(* Logix 5000 project; controller PLC_MCC1300_75F1 vendor 1 type 14 code 166 rev 32.11; software revision 32.04; part 44 of 83 *)
(* tags used below, declared in another part *)
   CONST_tPlant : UDT_PLANT_CONSTANTS;
   GP_OB_InitializeMain : GP_OB_Initialize;
   GP_PosWindow : GP_PosWindow;
   GP_TrackingSearchPlate : GP_TrackingSearchPlate;
   M307ASpeedUp : MAC_SpeedUp;
   M307ASpeedUp_ALM : MAC_SpeedUp_ALM;
   M30xTrimDeck : MAC_TrimmingDeck[5];
   M30xTrimDeck_ALM : MAC_TrimmingDeck_ALM[5];
   M30xTrimDeck_HMR : MAC_TrimmingDeck_HMR[5];
   TMP_d : DINT;
   TMP_dIndex : DINT;
   TMP_dIndexMotor : DINT;
   TMP_dLineSpeed : DINT;
   TMP_r : REAL;
   TMP_x : BOOL;
   xAlwaysOFF : BOOL;
   xDebugOFF : BOOL;
   Z200_SnapDataEth : UDT_ConvoyCap_ZC[2];
   Z300_BufferPlate : UDT_LINE_BUFFER_PLATE;
   Z300_Conveyor : UDT_StandConv[29];
   Z300_LineTracking : UDT_LINE_TRACKING;
   Z301 : MAC_Zone_ML;
   Z301_HMR : MAC_Zone_ML_HMR;
   Z301_HMW : MAC_Zone_ML_HMW;
(* MainProgram, continued *)

ROUTINE M307ASpeedUp_Faults   (* ladder *)
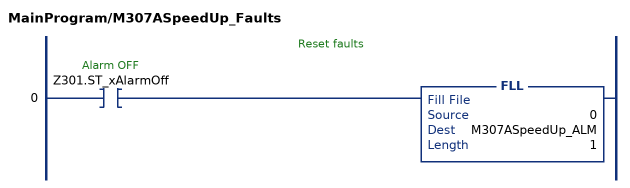
   // Reset faults
   0: XIC(Z301.ST_xAlarmOff)FLL(0,M307ASpeedUp_ALM,1);
END_ROUTINE

ROUTINE M307ASpeedUp_Logic   (* ladder *)
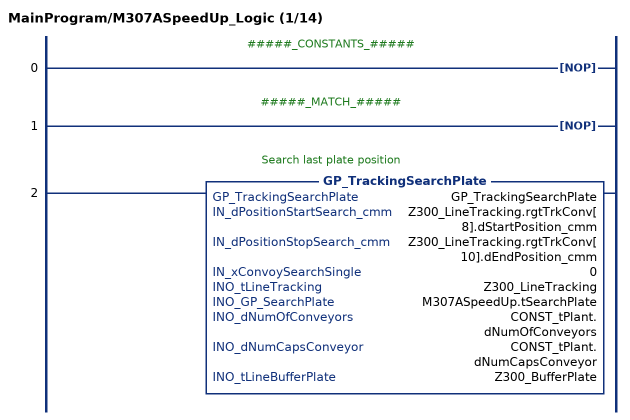
   // #####_CONSTANTS_#####
   0: NOP();
   // #####_MATCH_#####
   1: NOP();
   // Search last plate position
   2: GP_TrackingSearchPlate(GP_TrackingSearchPlate,Z300_LineTracking.rgtTrkConv[8].dStartPosition_cmm,Z300_LineTracking.rgtTrkConv[10].dEndPosition_cmm,0,Z300_LineTracking,M307ASpeedUp.tSearchPlate,CONST_tPlant.dNumOfConveyors,CONST_tPlant.dNumCapsConveyor,Z300_BufferPlate);
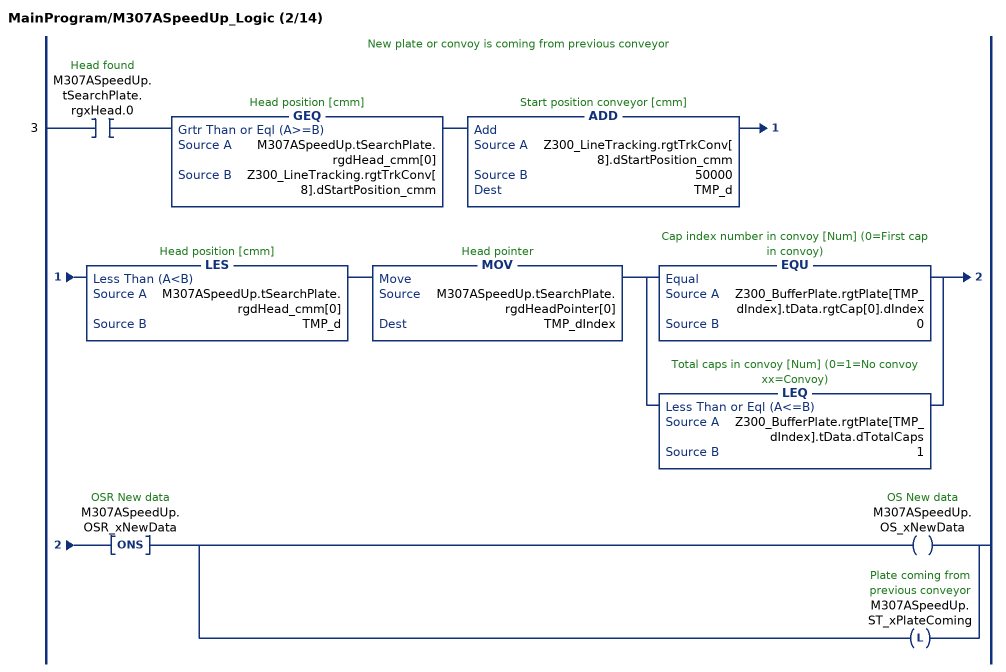
   // New plate or convoy is coming from previous conveyor
   3: XIC(M307ASpeedUp.tSearchPlate.rgxHead.0)GEQ(M307ASpeedUp.tSearchPlate.rgdHead_cmm[0],Z300_LineTracking.rgtTrkConv[8].dStartPosition_cmm)ADD(Z300_LineTracking.rgtTrkConv[8].dStartPosition_cmm,50000,TMP_d)LES(M307ASpeedUp.tSearchPlate.rgdHead_cmm[0],TMP_d)MOV(M307ASpeedUp.tSearchPlate.rgdHeadPointer[0],TMP_dIndex)[EQU(Z300_BufferPlate.rgtPlate[TMP_dIndex].tData.rgtCap[0].dIndex,0) ,LEQ(Z300_BufferPlate.rgtPlate[TMP_dIndex].tData.dTotalCaps,1) ]ONS(M307ASpeedUp.OSR_xNewData)[OTE(M307ASpeedUp.OS_xNewData) ,OTL(M307ASpeedUp.ST_xPlateComing) ];
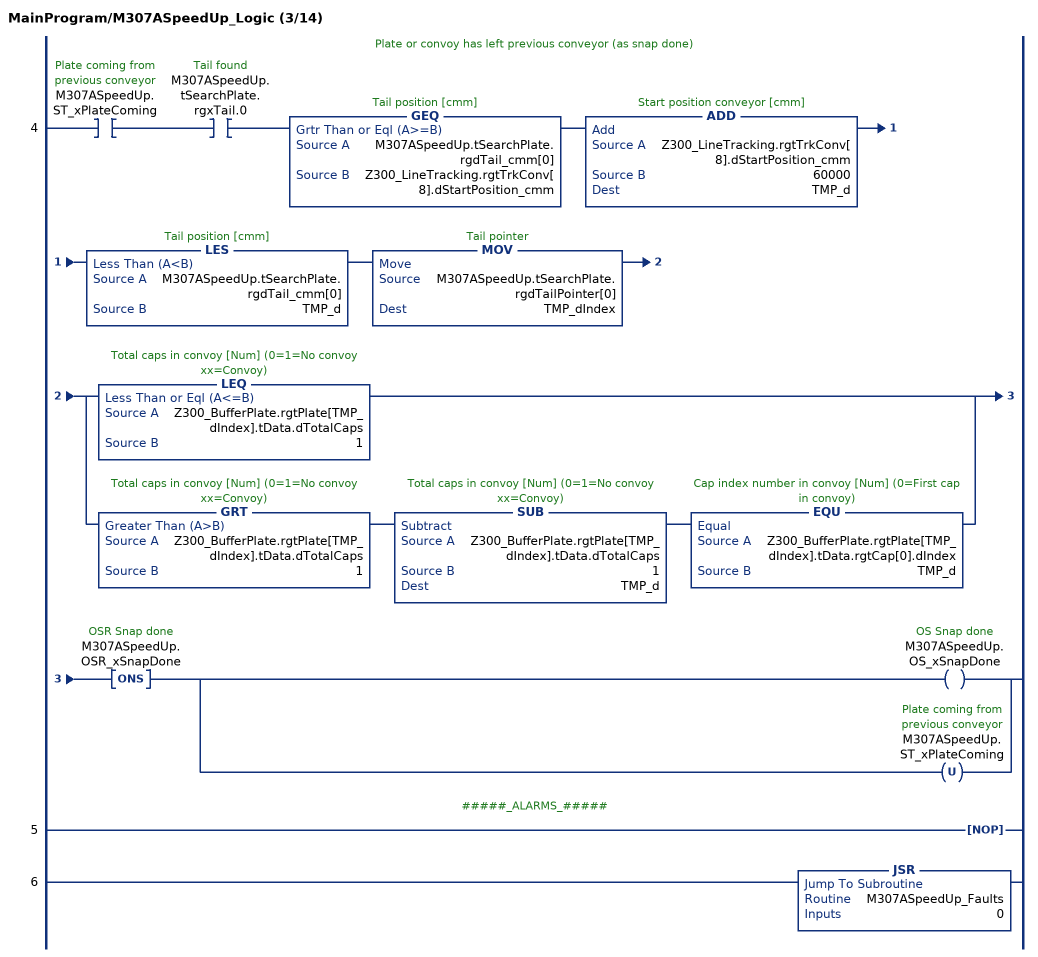
   // Plate or convoy has left previous conveyor (as snap done)
   4: XIC(M307ASpeedUp.ST_xPlateComing)XIC(M307ASpeedUp.tSearchPlate.rgxTail.0)GEQ(M307ASpeedUp.tSearchPlate.rgdTail_cmm[0],Z300_LineTracking.rgtTrkConv[8].dStartPosition_cmm)ADD(Z300_LineTracking.rgtTrkConv[8].dStartPosition_cmm,60000,TMP_d)LES(M307ASpeedUp.tSearchPlate.rgdTail_cmm[0],TMP_d)MOV(M307ASpeedUp.tSearchPlate.rgdTailPointer[0],TMP_dIndex)[LEQ(Z300_BufferPlate.rgtPlate[TMP_dIndex].tData.dTotalCaps,1) ,GRT(Z300_BufferPlate.rgtPlate[TMP_dIndex].tData.dTotalCaps,1) SUB(Z300_BufferPlate.rgtPlate[TMP_dIndex].tData.dTotalCaps,1,TMP_d) EQU(Z300_BufferPlate.rgtPlate[TMP_dIndex].tData.rgtCap[0].dIndex,TMP_d) ]ONS(M307ASpeedUp.OSR_xSnapDone)[OTE(M307ASpeedUp.OS_xSnapDone) ,OTU(M307ASpeedUp.ST_xPlateComing) ];
   // #####_ALARMS_#####
   5: NOP();
   6: JSR(M307ASpeedUp_Faults,0);
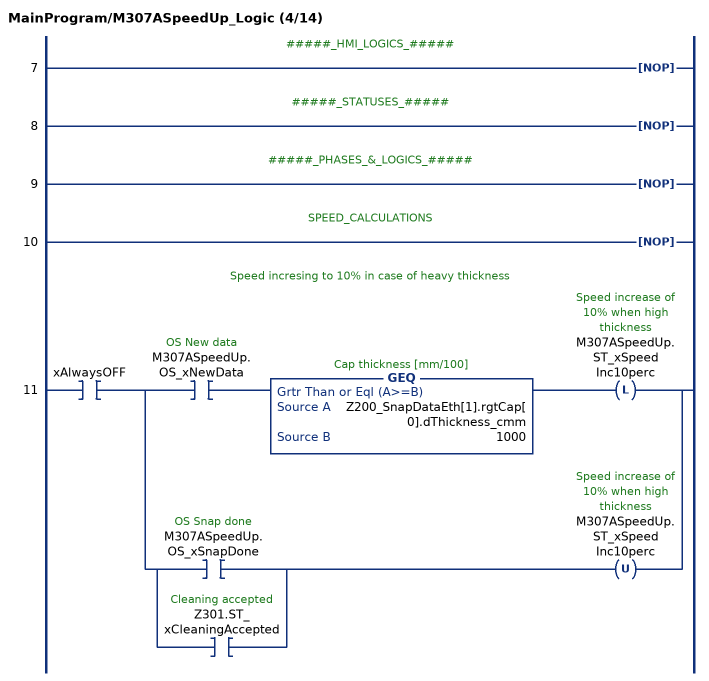
   // #####_HMI_LOGICS_#####
   7: NOP();
   // #####_STATUSES_#####
   8: NOP();
   // #####_PHASES_&_LOGICS_#####
   9: NOP();
   // SPEED_CALCULATIONS
   10: NOP();
   // Speed incresing to 10% in case of heavy thickness
   11: XIC(xAlwaysOFF)[XIC(M307ASpeedUp.OS_xNewData) GEQ(Z200_SnapDataEth[1].rgtCap[0].dThickness_cmm,1000) OTL(M307ASpeedUp.ST_xSpeedInc10perc) ,[XIC(M307ASpeedUp.OS_xSnapDone) ,XIC(Z301.ST_xCleaningAccepted) ] OTU(M307ASpeedUp.ST_xSpeedInc10perc) ];
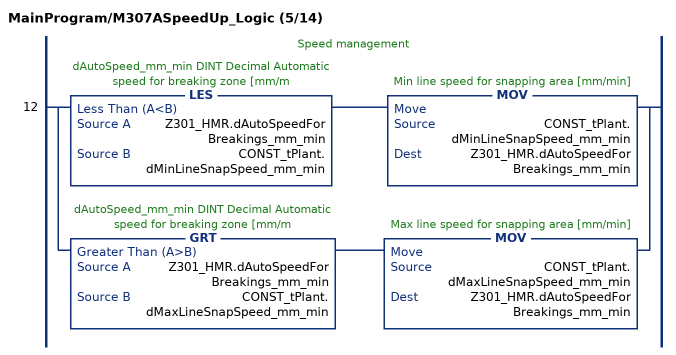
   // Speed management
   12: [LES(Z301_HMR.dAutoSpeedForBreakings_mm_min,CONST_tPlant.dMinLineSnapSpeed_mm_min) MOV(CONST_tPlant.dMinLineSnapSpeed_mm_min,Z301_HMR.dAutoSpeedForBreakings_mm_min) ,GRT(Z301_HMR.dAutoSpeedForBreakings_mm_min,CONST_tPlant.dMaxLineSnapSpeed_mm_min) MOV(CONST_tPlant.dMaxLineSnapSpeed_mm_min,Z301_HMR.dAutoSpeedForBreakings_mm_min) ];
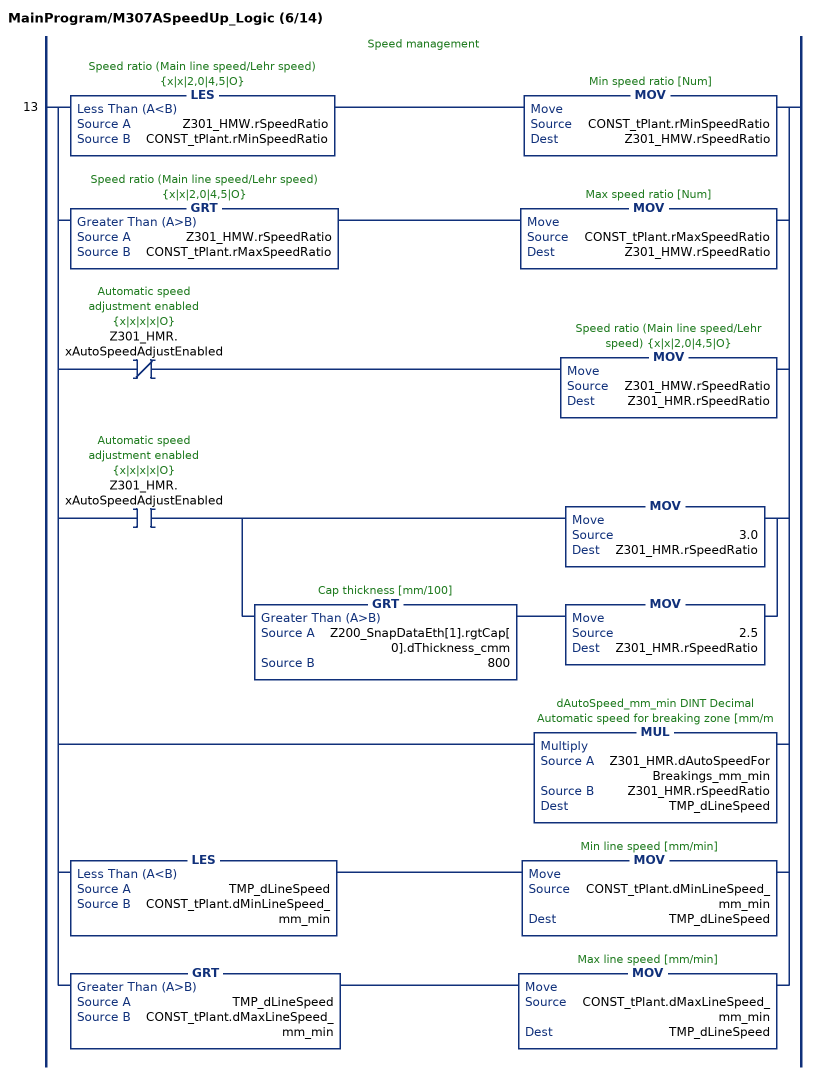
   // Speed management
   13: [LES(Z301_HMW.rSpeedRatio,CONST_tPlant.rMinSpeedRatio) MOV(CONST_tPlant.rMinSpeedRatio,Z301_HMW.rSpeedRatio) ,GRT(Z301_HMW.rSpeedRatio,CONST_tPlant.rMaxSpeedRatio) MOV(CONST_tPlant.rMaxSpeedRatio,Z301_HMW.rSpeedRatio) ,XIO(Z301_HMR.xAutoSpeedAdjustEnabled) MOV(Z301_HMW.rSpeedRatio,Z301_HMR.rSpeedRatio) ,XIC(Z301_HMR.xAutoSpeedAdjustEnabled) [MOV(3.0,Z301_HMR.rSpeedRatio) ,GRT(Z200_SnapDataEth[1].rgtCap[0].dThickness_cmm,800) MOV(2.5,Z301_HMR.rSpeedRatio) ] ,MUL(Z301_HMR.dAutoSpeedForBreakings_mm_min,Z301_HMR.rSpeedRatio,TMP_dLineSpeed) ,LES(TMP_dLineSpeed,CONST_tPlant.dMinLineSpeed_mm_min) MOV(CONST_tPlant.dMinLineSpeed_mm_min,TMP_dLineSpeed) ,GRT(TMP_dLineSpeed,CONST_tPlant.dMaxLineSpeed_mm_min) MOV(CONST_tPlant.dMaxLineSpeed_mm_min,TMP_dLineSpeed) ];
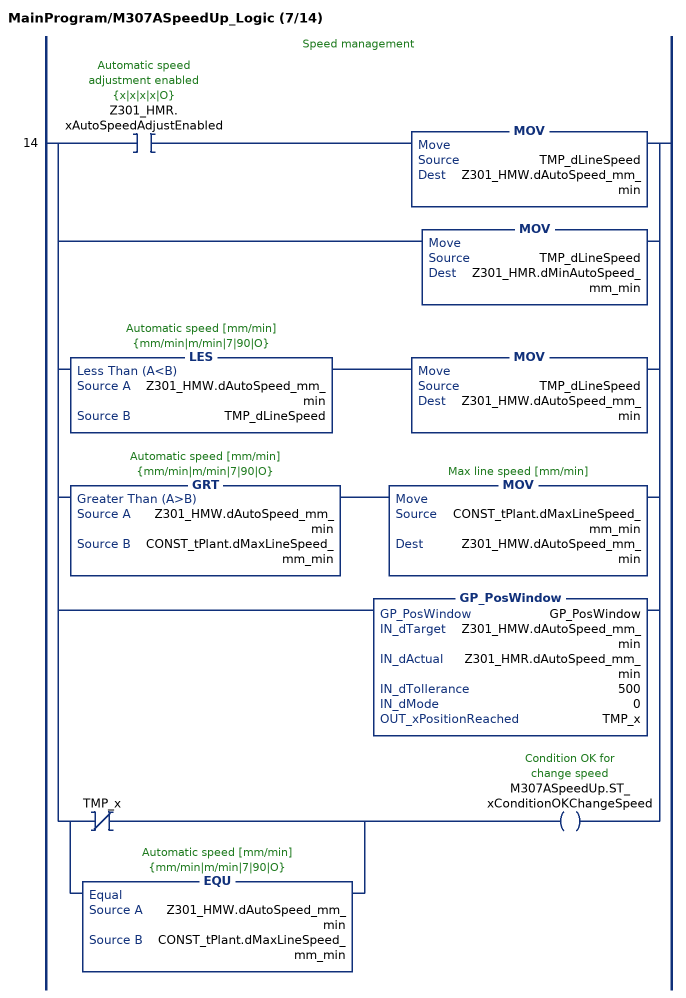
   // Speed management
   14: [XIC(Z301_HMR.xAutoSpeedAdjustEnabled) MOV(TMP_dLineSpeed,Z301_HMW.dAutoSpeed_mm_min) ,MOV(TMP_dLineSpeed,Z301_HMR.dMinAutoSpeed_mm_min) ,LES(Z301_HMW.dAutoSpeed_mm_min,TMP_dLineSpeed) MOV(TMP_dLineSpeed,Z301_HMW.dAutoSpeed_mm_min) ,GRT(Z301_HMW.dAutoSpeed_mm_min,CONST_tPlant.dMaxLineSpeed_mm_min) MOV(CONST_tPlant.dMaxLineSpeed_mm_min,Z301_HMW.dAutoSpeed_mm_min) ,[GP_PosWindow(GP_PosWindow,Z301_HMW.dAutoSpeed_mm_min,Z301_HMR.dAutoSpeed_mm_min,500,0,TMP_x) ,[XIO(TMP_x) ,EQU(Z301_HMW.dAutoSpeed_mm_min,CONST_tPlant.dMaxLineSpeed_mm_min) ] OTE(M307ASpeedUp.ST_xConditionOKChangeSpeed) ] ];
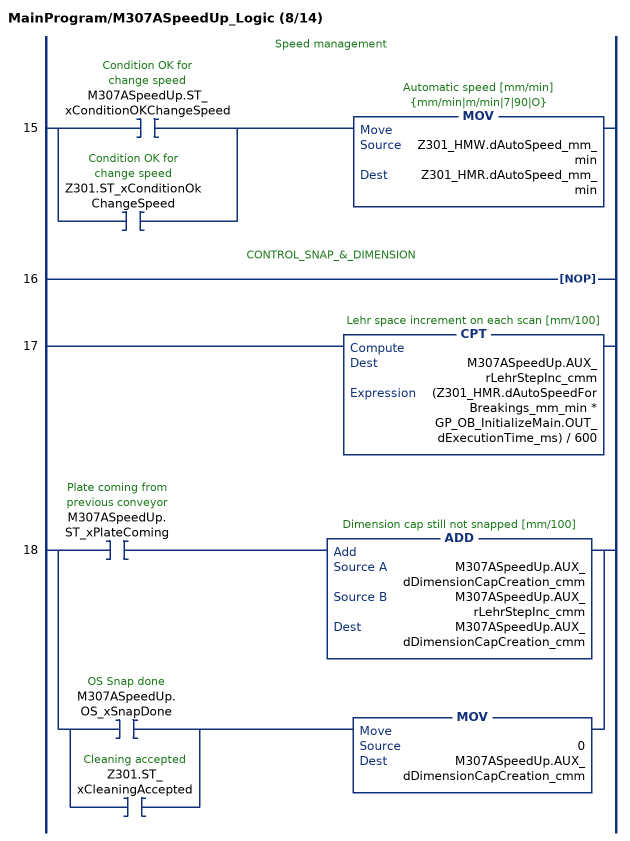
   // Speed management
   15: [XIC(M307ASpeedUp.ST_xConditionOKChangeSpeed) ,XIC(Z301.ST_xConditionOkChangeSpeed) ]MOV(Z301_HMW.dAutoSpeed_mm_min,Z301_HMR.dAutoSpeed_mm_min);
   // CONTROL_SNAP_&_DIMENSION
   16: NOP();
   17: CPT(M307ASpeedUp.AUX_rLehrStepInc_cmm,(Z301_HMR.dAutoSpeedForBreakings_mm_min * GP_OB_InitializeMain.OUT_dExecutionTime_ms) / 600);
   18: [XIC(M307ASpeedUp.ST_xPlateComing) ADD(M307ASpeedUp.AUX_dDimensionCapCreation_cmm,M307ASpeedUp.AUX_rLehrStepInc_cmm,M307ASpeedUp.AUX_dDimensionCapCreation_cmm) ,[XIC(M307ASpeedUp.OS_xSnapDone) ,XIC(Z301.ST_xCleaningAccepted) ] MOV(0,M307ASpeedUp.AUX_dDimensionCapCreation_cmm) ];
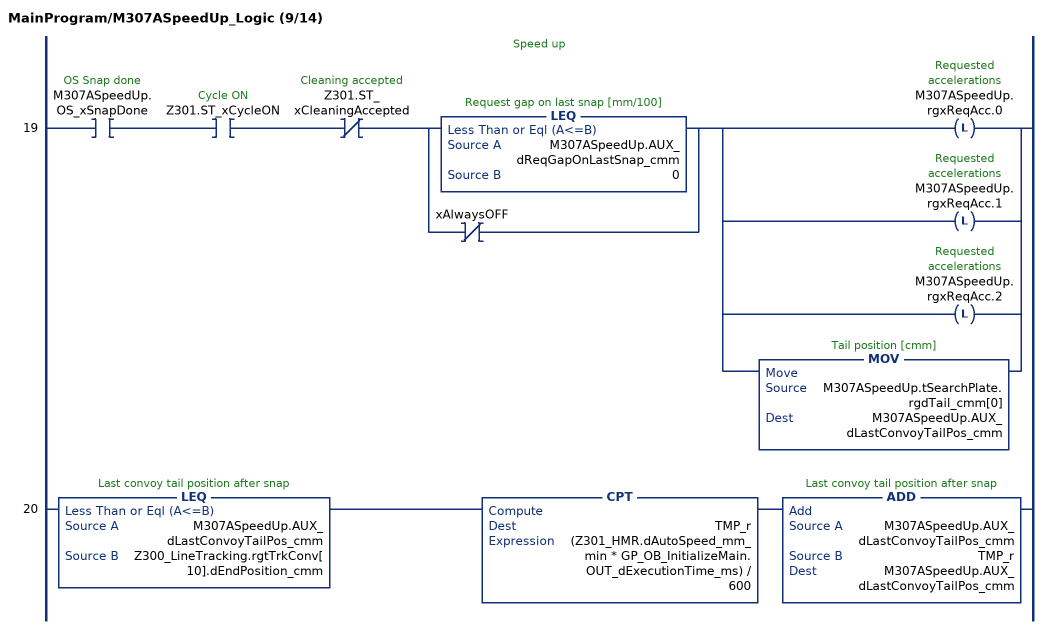
   // Speed up
   19: XIC(M307ASpeedUp.OS_xSnapDone)XIC(Z301.ST_xCycleON)XIO(Z301.ST_xCleaningAccepted)[LEQ(M307ASpeedUp.AUX_dReqGapOnLastSnap_cmm,0) ,XIO(xAlwaysOFF) ][OTL(M307ASpeedUp.rgxReqAcc.0) ,OTL(M307ASpeedUp.rgxReqAcc.1) ,OTL(M307ASpeedUp.rgxReqAcc.2) ,MOV(M307ASpeedUp.tSearchPlate.rgdTail_cmm[0],M307ASpeedUp.AUX_dLastConvoyTailPos_cmm) ];
   20: LEQ(M307ASpeedUp.AUX_dLastConvoyTailPos_cmm,Z300_LineTracking.rgtTrkConv[10].dEndPosition_cmm)CPT(TMP_r,(Z301_HMR.dAutoSpeed_mm_min * GP_OB_InitializeMain.OUT_dExecutionTime_ms) / 600)ADD(M307ASpeedUp.AUX_dLastConvoyTailPos_cmm,TMP_r,M307ASpeedUp.AUX_dLastConvoyTailPos_cmm);
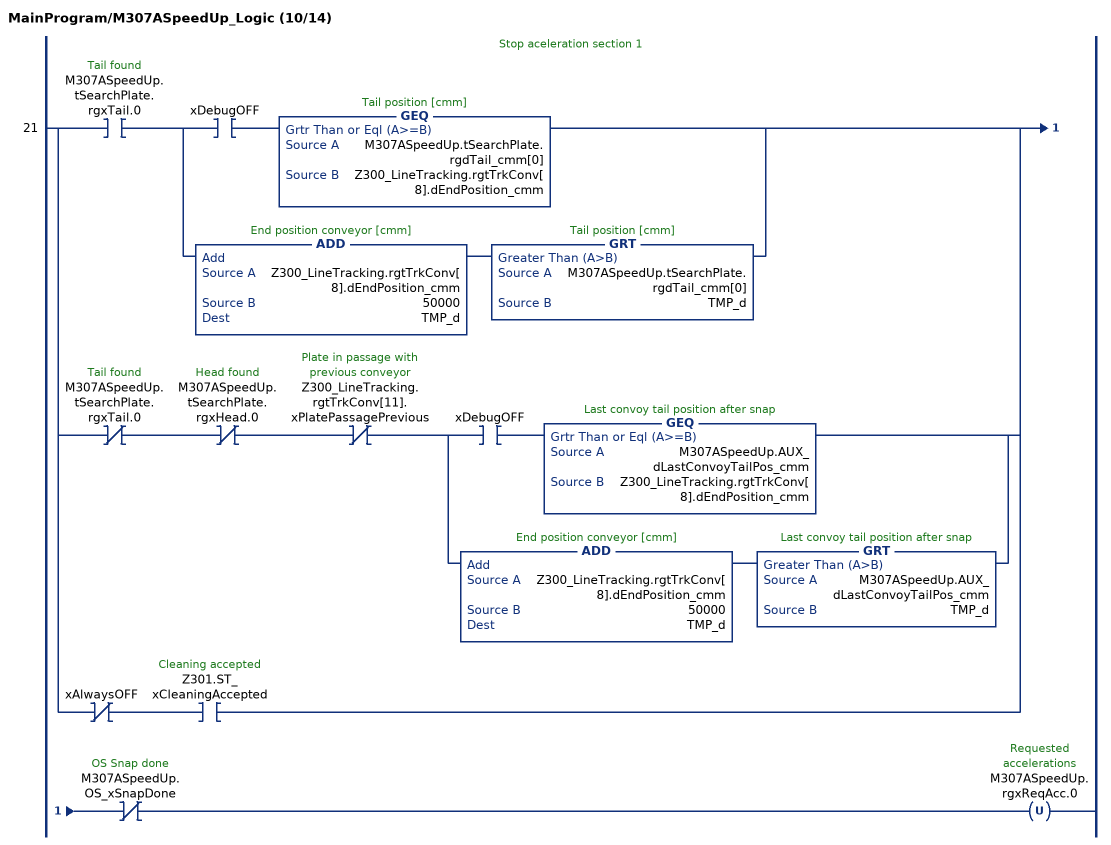
   // Stop aceleration section 1
   21: [XIC(M307ASpeedUp.tSearchPlate.rgxTail.0) [XIC(xDebugOFF) GEQ(M307ASpeedUp.tSearchPlate.rgdTail_cmm[0],Z300_LineTracking.rgtTrkConv[8].dEndPosition_cmm) ,ADD(Z300_LineTracking.rgtTrkConv[8].dEndPosition_cmm,50000,TMP_d) GRT(M307ASpeedUp.tSearchPlate.rgdTail_cmm[0],TMP_d) ] ,XIO(M307ASpeedUp.tSearchPlate.rgxTail.0) XIO(M307ASpeedUp.tSearchPlate.rgxHead.0) XIO(Z300_LineTracking.rgtTrkConv[11].xPlatePassagePrevious) [XIC(xDebugOFF) GEQ(M307ASpeedUp.AUX_dLastConvoyTailPos_cmm,Z300_LineTracking.rgtTrkConv[8].dEndPosition_cmm) ,ADD(Z300_LineTracking.rgtTrkConv[8].dEndPosition_cmm,50000,TMP_d) GRT(M307ASpeedUp.AUX_dLastConvoyTailPos_cmm,TMP_d) ] ,XIO(xAlwaysOFF) XIC(Z301.ST_xCleaningAccepted) ]XIO(M307ASpeedUp.OS_xSnapDone)OTU(M307ASpeedUp.rgxReqAcc.0);
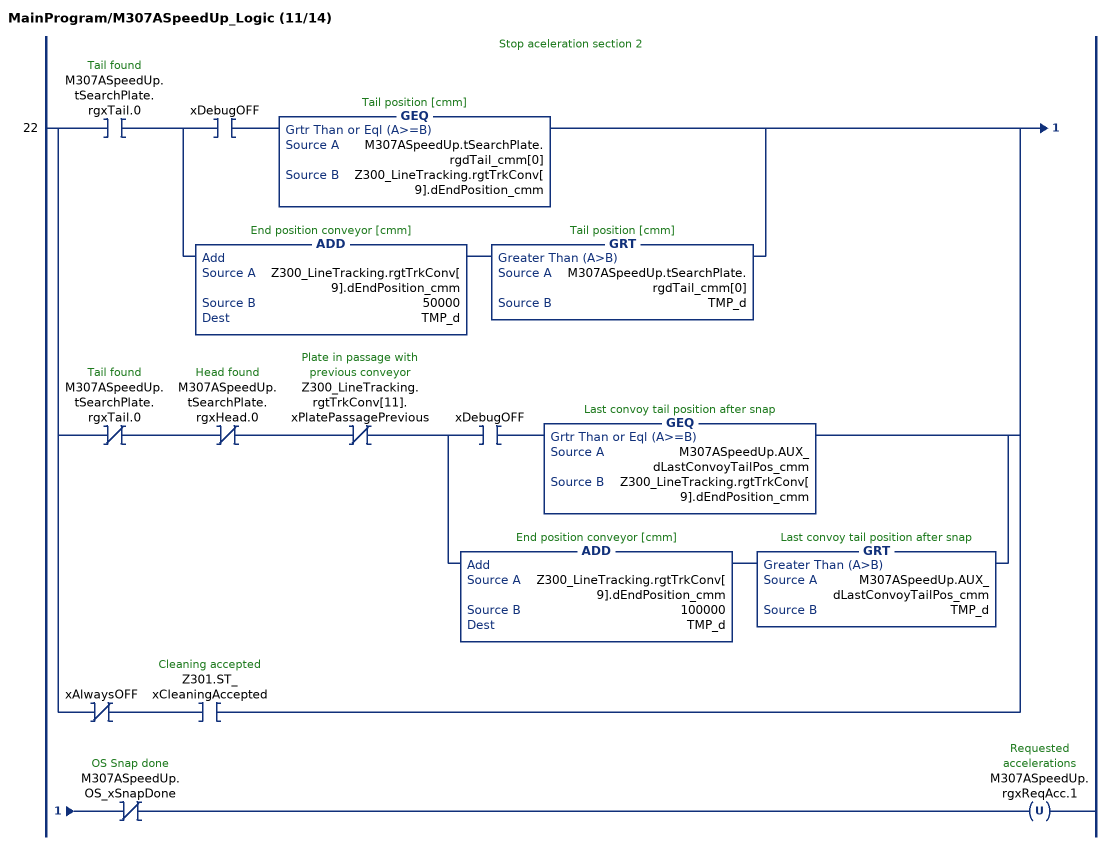
   // Stop aceleration section 2
   22: [XIC(M307ASpeedUp.tSearchPlate.rgxTail.0) [XIC(xDebugOFF) GEQ(M307ASpeedUp.tSearchPlate.rgdTail_cmm[0],Z300_LineTracking.rgtTrkConv[9].dEndPosition_cmm) ,ADD(Z300_LineTracking.rgtTrkConv[9].dEndPosition_cmm,50000,TMP_d) GRT(M307ASpeedUp.tSearchPlate.rgdTail_cmm[0],TMP_d) ] ,XIO(M307ASpeedUp.tSearchPlate.rgxTail.0) XIO(M307ASpeedUp.tSearchPlate.rgxHead.0) XIO(Z300_LineTracking.rgtTrkConv[11].xPlatePassagePrevious) [XIC(xDebugOFF) GEQ(M307ASpeedUp.AUX_dLastConvoyTailPos_cmm,Z300_LineTracking.rgtTrkConv[9].dEndPosition_cmm) ,ADD(Z300_LineTracking.rgtTrkConv[9].dEndPosition_cmm,100000,TMP_d) GRT(M307ASpeedUp.AUX_dLastConvoyTailPos_cmm,TMP_d) ] ,XIO(xAlwaysOFF) XIC(Z301.ST_xCleaningAccepted) ]XIO(M307ASpeedUp.OS_xSnapDone)OTU(M307ASpeedUp.rgxReqAcc.1);